
screen "716_TS_IF_NOT_USED" 1280x800, template "Top_Header"
   on GenerateScreen: "SDC_TS_REFERENCE"("SDC\_TS_Nr"); "SDC_TS_IF"(); SetTag("DB_SDC_TS_IF_HMI.HMI[XX].BILD_Nr", 716); SetTag("SDC\_intern_Bildnummer", 716)
   on ClearScreen: SetTag("DB_SDC_TS_IF_HMI.HMI[XX].BILD_Nr", 0)
   TextField "Textfeld_18" at 739,287 size 178x25; Text 'acknowledge error / Command forward'
   Circle "Kreis_27" at 716,292 size 15x15
      Appearance <- "DB_SDC_TS_IF_COMMAND.SEK[XXX].BIT1"
   TextField "Textfeld_1" at 739,304 size 191x25; Text '1 = automatic in section / Command forward'
   Circle "Kreis_1" at 716,308 size 15x15
      Appearance <- "DB_SDC_TS_IF_COMMAND.SEK[XXX].BIT1"
   TextField "Textfeld_2" at 739,319 size 202x25; Text '1 = manual in section / Command forward'
   Circle "Kreis_2" at 716,324 size 15x15
      Appearance <- "DB_SDC_TS_IF_COMMAND.SEK[XXX].BIT1"
   TextField "Textfeld_4" at 739,336 size 201x25; Text 'spare / Command forward / Spare'
   Circle "Kreis_3" at 716,340 size 15x15
      Appearance <- "DB_SDC_TS_IF_COMMAND.SEK[XXX].BIT1"
   TextField "Textfeld_5" at 955,286 size 194x25; Text 'spare / Command forward / Spare'
   Circle "Kreis_4" at 932,291 size 15x15
      Appearance <- "DB_SDC_TS_IF_COMMAND.SEK[XXX].BIT1"
   TextField "Textfeld_6" at 955,303 size 150x25; Text '1 = emergency stop / Command forward'
   Circle "Kreis_5" at 932,307 size 15x15
      Appearance <- "DB_SDC_TS_IF_COMMAND.SEK[XXX].BIT1"
   TextField "Textfeld_7" at 955,318 size 138x25; Text 'spare / Command forward / Spare'
   Circle "Kreis_6" at 932,323 size 15x15
      Appearance <- "DB_SDC_TS_IF_COMMAND.SEK[XXX].BIT1"
   TextField "Textfeld_9" at 738,389 size 125x22; Text 'forward / Command forward'
   Circle "Kreis_8" at 715,394 size 15x15
      Appearance <- "DB_SDC_TS_IF_COMMAND.SEK[XXX].BIT1"
   TextField "Textfeld_10" at 738,406 size 125x22; Text 'backward / Command forward'
   Circle "Kreis_9" at 715,410 size 15x15
      Appearance <- "DB_SDC_TS_IF_COMMAND.SEK[XXX].BIT1"
   TextField "Textfeld_11" at 738,421 size 136x22; Text 'bypass stop position / Command forward'
   Circle "Kreis_10" at 715,426 size 15x15
      Appearance <- "DB_SDC_TS_IF_COMMAND.SEK[XXX].BIT1"
   TextField "Textfeld_12" at 738,438 size 125x22; Text 'speed setpoint 1 / Command forward / Speed Setpoint 1'
   Circle "Kreis_11" at 715,442 size 15x15
      Appearance <- "DB_SDC_TS_IF_COMMAND.SEK[XXX].BIT1"
   TextField "Textfeld_13" at 738,453 size 125x22; Text 'speed setpoint 2 / Command forward / Speed Setpoint 2'
   Circle "Kreis_12" at 715,458 size 15x15
      Appearance <- "DB_SDC_TS_IF_COMMAND.SEK[XXX].BIT1"
   TextField "Textfeld_14" at 738,470 size 156x22; Text 'variable speed setpoint / Command forward / Variable Speed Setpoint'
   Circle "Kreis_13" at 715,474 size 15x15
      Appearance <- "DB_SDC_TS_IF_COMMAND.SEK[XXX].BIT1"
   TextField "Textfeld_15" at 738,485 size 179x22; Text 'enable before stop position / Command forward'
   Circle "Kreis_14" at 715,490 size 15x15
      Appearance <- "DB_SDC_TS_IF_COMMAND.SEK[XXX].BIT1"
   TextField "Textfeld_16" at 738,502 size 168x22; Text 'enable after stop position / Command forward'
   Circle "Kreis_15" at 715,506 size 15x15
      Appearance <- "DB_SDC_TS_IF_COMMAND.SEK[XXX].BIT1"
   TextField "Textfeld_17" at 894,187 size 170x27; Text 'commands / EMS-Number'
   TextField "Textfeld_19" at 625,407 size 27x114; Text 'bits / EMS-Number'
   IOField "EA-Feld_4" at 305,148 size 56x32; FormatPattern 9999
      on OnFinishInput: "SDC_TS_REFERENCE"("SDC\_TS_Nr"); "SDC_TS_IF"()
      ProcessValue <- "SDC\_TS_Nr"
   TextField "Textfeld_3" at 429,151 size 117x23; Text 'section no. / Sektionnumber / Section Number'
   Button "Schaltfläche_1" at 362,148 size 40x32; TextOff '+'
      on Click: function_dd21b452("SDC\_TS_Nr", 1); "SDC_TS_REFERENCE"("SDC\_TS_Nr"); "SDC_TS_IF"()
   Button "Schaltfläche_3" at 265,148 size 39x32; TextOff '-'
      on Click: function_b9b71300("SDC\_TS_Nr", 1); "SDC_TS_REFERENCE"("SDC\_TS_Nr"); "SDC_TS_IF"()
   IOField "EA-Feld_13" at 665,152 size 163x24; Authorization "Benutzerverwaltung"; FormatPattern ????????????????
      Appearance <- "SDC\DB_SDC_TS_PARAMETER\DB_SDC_TS_PARAMETER_HMI.HMI[XX].FR_EDIT"
      ProcessValue <- "SDC\DB_SDC_TS_REFERENCE\DB_SDC_TS_REFERENCE_X.Reference[XXX].Sektion"
      ObjectEnable <- "SDC\DB_SDC_TS_PARAMETER\DB_SDC_TS_PARAMETER_HMI.HMI[XX].FR_EDIT"
   TextField "Textfeld_20" at 625,218 size 27x114; Text 'values / EMS-Number / Values'
   IOField "EA-Feld_1" at 716,221 size 56x28; FormatPattern 99
      on OnFinishInput: "SDC_TS_PARAMETER"(); "SDC_TS_REFERENCE"("SDC\_TS_Nr")
      ProcessValue <- "DB_SDC_TS_IF_COMMAND.SEK[XXX].VAL.PROFIL"
   TextField "Textfeld_21" at 788,223 size 64x25; Text 'car type / Command forward'
   IOField "EA-Feld_2" at 716,237 size 56x28; FormatPattern 999999
      on OnFinishInput: "SDC_TS_PARAMETER"(); "SDC_TS_REFERENCE"("SDC\_TS_Nr")
      ProcessValue <- "DB_SDC_TS_IF_COMMAND.SEK[XXX].VAL.D_SETSPEED"
   TextField "Textfeld_22" at 788,239 size 202x25; Text 'setpoint drive speed mm/min / Command forward'
   IOField "EA-Feld_3" at 716,253 size 56x28; FormatPattern 99999
      on OnFinishInput: "SDC_TS_PARAMETER"(); "SDC_TS_REFERENCE"("SDC\_TS_Nr")
      ProcessValue <- "DB_SDC_TS_IF_COMMAND.SEK[XXX].VAL.D_POS_OFFS"
   TextField "Textfeld_23" at 788,255 size 192x25; Text 'stop position offset mm / Command forward / Stop positions offset mm'
   TextField "Textfeld_24" at 719,369 size 155x22; Text 'drive / Command forward'
   TextField "Textfeld_47" at 738,517 size 166x22; Text 'bypass distance controlle / Command forward / bypass distance control'
   Circle "Kreis_37" at 715,522 size 15x15
      Appearance <- "DB_SDC_TS_IF_COMMAND.SEK[XXX].BIT2"
   TextField "Textfeld_48" at 955,335 size 84x25; Text 'set car type / Command forward'
   Circle "Kreis_38" at 932,339 size 15x15
      Appearance <- "DB_SDC_TS_IF_COMMAND.SEK[XXX].BIT2"
   TextField "Textfeld_49" at 625,657 size 27x59; Text 'fkt / EMS-Number'
   TextField "Textfeld_50" at 766,592 size 155x22; Text 'set / Command forward / Set'
   TextField "Textfeld_51" at 738,612 size 143x22; Text 'EMS to maintenace 1 / Command forward'
   Circle "Kreis_39" at 715,617 size 15x15
      Appearance <- "DB_SDC_TS_IF_COMMAND.SEK[XXX].FKT_SET"
   TextField "Textfeld_52" at 738,629 size 143x22; Text 'EMS to maintenace 2 / Command forward'
   Circle "Kreis_40" at 715,633 size 15x15
      Appearance <- "DB_SDC_TS_IF_COMMAND.SEK[XXX].FKT_SET"
   TextField "Textfeld_53" at 738,644 size 179x22; Text 'emerg. mode without hoist / Command forward'
   Circle "Kreis_41" at 715,649 size 15x15
      Appearance <- "DB_SDC_TS_IF_COMMAND.SEK[XXX].FKT_SET"
   TextField "Textfeld_55" at 738,660 size 129x22; Text 'emerg. mode drive / Command forward'
   Circle "Kreis_43" at 715,665 size 15x15
      Appearance <- "DB_SDC_TS_IF_COMMAND.SEK[XXX].FKT_SET"
   TextField "Textfeld_57" at 738,684 size 125x22; Text 'PE check fault / Command forward / PE Check Fault'
   Circle "Kreis_45" at 715,689 size 15x15
      Appearance <- "DB_SDC_TS_IF_COMMAND.SEK[XXX].FKT_SET"
   TextField "Textfeld_58" at 738,701 size 125x22; Text 'brush check fault / Command forward'
   Circle "Kreis_46" at 715,705 size 15x15
      Appearance <- "DB_SDC_TS_IF_COMMAND.SEK[XXX].FKT_SET"
   TextField "Textfeld_59" at 1054,592 size 155x22; Text 'reset / Command forward / Reset'
   TextField "Textfeld_60" at 1026,612 size 143x22; Text 'EMS to maintenace 1 / Command forward'
   Circle "Kreis_47" at 1003,617 size 15x15
      Appearance <- "DB_SDC_TS_IF_COMMAND.SEK[XXX].FKT_RESET"
   TextField "Textfeld_61" at 1026,629 size 143x22; Text 'EMS to maintenace 2 / Command forward'
   Circle "Kreis_48" at 1003,633 size 15x15
      Appearance <- "DB_SDC_TS_IF_COMMAND.SEK[XXX].FKT_RESET"
   TextField "Textfeld_62" at 1026,644 size 179x22; Text 'emerg. mode without hoist / Command forward'
   Circle "Kreis_49" at 1003,649 size 15x15
      Appearance <- "DB_SDC_TS_IF_COMMAND.SEK[XXX].FKT_RESET"
   TextField "Textfeld_64" at 1026,660 size 129x22; Text 'emerg. mode drive / Command forward'
   Circle "Kreis_51" at 1003,665 size 15x15
      Appearance <- "DB_SDC_TS_IF_COMMAND.SEK[XXX].FKT_RESET"
   TextField "Textfeld_66" at 1026,684 size 125x22; Text 'PE check fault / Command forward / PE Check Fault'
   Circle "Kreis_53" at 1003,689 size 15x15
      Appearance <- "DB_SDC_TS_IF_COMMAND.SEK[XXX].FKT_RESET"
   TextField "Textfeld_67" at 1026,701 size 125x22; Text 'brush check fault / Command forward'
   Circle "Kreis_54" at 1003,705 size 15x15
      Appearance <- "DB_SDC_TS_IF_COMMAND.SEK[XXX].FKT_RESET"
   TextField "Textfeld_68" at 317,193 size 170x27; Text 'status / EMS-Number / Status'
   IOField "EA-Feld_5" at 169,212 size 56x28; FormatPattern 999
      on OnFinishInput: "SDC_TS_PARAMETER"(); "SDC_TS_REFERENCE"("SDC\_TS_Nr")
      ProcessValue <- "DB_SDC_TS_IF_STATUS.SEK[XXX].VAL.EMS_ID"
   TextField "Textfeld_69" at 225,215 size 60x25; Text 'EMS ID / Command forward'
   IOField "EA-Feld_6" at 169,228 size 56x28; FormatPattern 99
      on OnFinishInput: "SDC_TS_PARAMETER"(); "SDC_TS_REFERENCE"("SDC\_TS_Nr")
      ProcessValue <- "DB_SDC_TS_IF_STATUS.SEK[XXX].VAL.PROFIL"
   TextField "Textfeld_70" at 225,231 size 60x25; Text 'car type / Command forward'
   IOField "EA-Feld_7" at 139,244 size 86x28; FormatPattern 9999999999
      on OnFinishInput: "SDC_TS_PARAMETER"(); "SDC_TS_REFERENCE"("SDC\_TS_Nr")
      ProcessValue <- "DB_SDC_TS_IF_STATUS.SEK[XXX].VAL.DRIVE_POS"
   TextField "Textfeld_71" at 225,247 size 170x25; Text 'drive position mm / Command forward'
   IOField "EA-Feld_10" at 385,213 size 56x28; FormatPattern 999
      on OnFinishInput: "SDC_TS_PARAMETER"(); "SDC_TS_REFERENCE"("SDC\_TS_Nr")
      ProcessValue <- "DB_SDC_TS_IF_STATUS.SEK[XXX].VAL.ERROR"
   TextField "Textfeld_74" at 443,215 size 60x25; Text 'error no. / Command forward'
   IOField "EA-Feld_11" at 385,229 size 56x28; FormatPattern 999
      on OnFinishInput: "SDC_TS_PARAMETER"(); "SDC_TS_REFERENCE"("SDC\_TS_Nr")
      ProcessValue <- "DB_SDC_TS_IF_STATUS.SEK[XXX].VAL.DRIVE_POS_PERC"
   TextField "Textfeld_75" at 443,231 size 162x25; Text 'position in % at sektion / Command forward / Position in % in Sektion'
   IOField "EA-Feld_12" at 385,245 size 56x28; FormatPattern 999
      on OnFinishInput: "SDC_TS_PARAMETER"(); "SDC_TS_REFERENCE"("SDC\_TS_Nr")
      ProcessValue <- "DB_SDC_TS_IF_STATUS.SEK[XXX].VAL.SEK"
   TextField "Textfeld_76" at 443,247 size 162x25; Text 'sektion / Command forward / Section'
   TextField "Textfeld_77" at 179,287 size 178x25; Text 'EMS present / Command forward'
   Circle "Kreis_55" at 156,292 size 15x15
      Appearance <- "DB_SDC_TS_IF_STATUS.SEK[XXX].BIT1"
   TextField "Textfeld_78" at 179,304 size 191x25; Text 'general error / Command forward'
   Circle "Kreis_56" at 156,308 size 15x15
      Appearance <- "DB_SDC_TS_IF_STATUS.SEK[XXX].BIT1"
   TextField "Textfeld_79" at 179,319 size 202x25; Text 'EMS in manual mode (IR) / Command forward'
   Circle "Kreis_57" at 156,324 size 15x15
      Appearance <- "DB_SDC_TS_IF_STATUS.SEK[XXX].BIT1"
   TextField "Textfeld_80" at 179,336 size 201x25; Text 'more than 1 EMS in section / Command forward'
   Circle "Kreis_58" at 156,340 size 15x15
      Appearance <- "DB_SDC_TS_IF_STATUS.SEK[XXX].BIT1"
   TextField "Textfeld_81" at 395,286 size 194x25; Text 'error on commands / Command forward'
   Circle "Kreis_59" at 372,291 size 15x15
      Appearance <- "DB_SDC_TS_IF_STATUS.SEK[XXX].BIT1"
   TextField "Textfeld_82" at 395,303 size 229x25; Text 'warning distance controll / Command forward / "1" -> No Stop'
   Circle "Kreis_60" at 372,307 size 15x15
      Appearance <- "DB_SDC_TS_IF_STATUS.SEK[XXX].BIT1"
   TextField "Textfeld_83" at 395,318 size 138x25; Text 'spare / Command forward / Spare'
   Circle "Kreis_61" at 372,323 size 15x15
      Appearance <- "DB_SDC_TS_IF_STATUS.SEK[XXX].BIT1"
   TextField "Textfeld_84" at 395,335 size 220x25; Text 'error code is a warning / Command forward'
   Circle "Kreis_62" at 372,339 size 15x15
      Appearance <- "DB_SDC_TS_IF_STATUS.SEK[XXX].BIT1"
   TextField "Textfeld_85" at 163,369 size 155x22; Text 'drive / Command forward'
   TextField "Textfeld_88" at 186,389 size 125x22; Text 'drive is on / Command forward'
   Circle "Kreis_63" at 163,394 size 15x15
      Appearance <- "DB_SDC_TS_IF_STATUS.SEK[XXX].BIT1"
   TextField "Textfeld_89" at 186,406 size 125x22; Text 'drive is off / Command forward'
   Circle "Kreis_64" at 163,410 size 15x15
      Appearance <- "DB_SDC_TS_IF_STATUS.SEK[XXX].BIT1"
   TextField "Textfeld_94" at 186,421 size 125x22; Text 'in position / Command forward'
   Circle "Kreis_69" at 163,426 size 15x15
      Appearance <- "DB_SDC_TS_IF_STATUS.SEK[XXX].BIT2"
   TextField "Textfeld_95" at 186,437 size 125x22; Text 'before position / Command forward'
   Circle "Kreis_70" at 163,442 size 15x15
      Appearance <- "DB_SDC_TS_IF_STATUS.SEK[XXX].BIT2"
   TextField "Textfeld_96" at 186,453 size 125x22; Text 'after position / Command forward'
   Circle "Kreis_71" at 163,458 size 15x15
      Appearance <- "DB_SDC_TS_IF_STATUS.SEK[XXX].BIT2"
   TextField "Textfeld_97" at 186,469 size 125x22; Text 'after actionpoint 1 / Command forward'
   Circle "Kreis_72" at 163,474 size 15x15
      Appearance <- "DB_SDC_TS_IF_STATUS.SEK[XXX].BIT2"
   TextField "Textfeld_98" at 186,485 size 157x22; Text 'before/at actionpoint 1 / Command forward'
   Circle "Kreis_73" at 163,490 size 15x15
      Appearance <- "DB_SDC_TS_IF_STATUS.SEK[XXX].BIT2"
   TextField "Textfeld_99" at 186,501 size 125x22; Text 'after actionpoint 2 / Command forward'
   Circle "Kreis_74" at 163,506 size 15x15
      Appearance <- "DB_SDC_TS_IF_STATUS.SEK[XXX].BIT2"
   TextField "Textfeld_100" at 186,517 size 152x22; Text 'before/at actionpoint 2 / Command forward'
   Circle "Kreis_75" at 163,522 size 15x15
      Appearance <- "DB_SDC_TS_IF_STATUS.SEK[XXX].BIT2"
   TextField "Textfeld_133" at 186,533 size 125x22; Text 'forwards / Command forward'
   Circle "Kreis_108" at 163,538 size 15x15
      Appearance <- "DB_SDC_TS_IF_STATUS.SEK[XXX].BIT4"
   TextField "Textfeld_134" at 186,550 size 125x22; Text 'backwards / Command forward'
   Circle "Kreis_109" at 163,554 size 15x15
      Appearance <- "DB_SDC_TS_IF_STATUS.SEK[XXX].BIT4"
   TextField "Textfeld_38" at 738,717 size 176x22; Text 'communication check fault / Command forward'
   Circle "Kreis_29" at 715,721 size 15x15
      Appearance <- "DB_SDC_TS_IF_COMMAND.SEK[XXX].FKT_SET"
   TextField "Textfeld_39" at 1026,717 size 176x22; Text 'communication check fault / Command forward'
   Circle "Kreis_30" at 1003,721 size 15x15
      Appearance <- "DB_SDC_TS_IF_COMMAND.SEK[XXX].FKT_RESET"

screen "722_ERRORS_NOT_USED" 1280x800, template "Top_Header"
   on GenerateScreen: "SDC_ERRORS"("HMI_EMS_Nr"); SetTag("SDC\_intern_Bildnummer", 722)
   TextField "Textfeld_18" at 235,235 size 31x132; Text '601 602 603 604 605 606 607 608 Command forward 601'
   Circle "Kreis_27" at 212,238 size 15x15
      Appearance <- "DB_SDC_ERRORS.EMS[XXX].DRIVE_1"
   Circle "Kreis_1" at 212,254 size 15x15
      Appearance <- "DB_SDC_ERRORS.EMS[XXX].DRIVE_1"
   Circle "Kreis_2" at 212,270 size 15x15
      Appearance <- "DB_SDC_ERRORS.EMS[XXX].DRIVE_1"
   Circle "Kreis_3" at 212,286 size 15x15
      Appearance <- "DB_SDC_ERRORS.EMS[XXX].DRIVE_1"
   Circle "Kreis_4" at 212,302 size 15x15
      Appearance <- "DB_SDC_ERRORS.EMS[XXX].DRIVE_1"
   Circle "Kreis_5" at 212,318 size 15x15
      Appearance <- "DB_SDC_ERRORS.EMS[XXX].DRIVE_1"
   Circle "Kreis_6" at 212,334 size 15x15
      Appearance <- "DB_SDC_ERRORS.EMS[XXX].DRIVE_1"
   Circle "Kreis_7" at 212,350 size 15x15
      Appearance <- "DB_SDC_ERRORS.EMS[XXX].DRIVE_1"
   TextField "Textfeld_9" at 292,235 size 31x132; Text '609 610 611 612 613 614 615 616 Command forward 609'
   Circle "Kreis_8" at 269,238 size 15x15
      Appearance <- "DB_SDC_ERRORS.EMS[XXX].DRIVE_1"
   Circle "Kreis_9" at 269,254 size 15x15
      Appearance <- "DB_SDC_ERRORS.EMS[XXX].DRIVE_1"
   Circle "Kreis_10" at 269,270 size 15x15
      Appearance <- "DB_SDC_ERRORS.EMS[XXX].DRIVE_1"
   Circle "Kreis_11" at 269,286 size 15x15
      Appearance <- "DB_SDC_ERRORS.EMS[XXX].DRIVE_1"
   Circle "Kreis_12" at 269,302 size 15x15
      Appearance <- "DB_SDC_ERRORS.EMS[XXX].DRIVE_1"
   Circle "Kreis_13" at 269,318 size 15x15
      Appearance <- "DB_SDC_ERRORS.EMS[XXX].DRIVE_1"
   Circle "Kreis_14" at 269,334 size 15x15
      Appearance <- "DB_SDC_ERRORS.EMS[XXX].DRIVE_1"
   Circle "Kreis_15" at 269,350 size 15x15
      Appearance <- "DB_SDC_ERRORS.EMS[XXX].DRIVE_1"
   TextField "Textfeld_17" at 271,202 size 100x38; Text 'drive / EMS-Number / Drive'
   TextField "Textfeld_19" at 180,241 size 32x114; Text 'generally / EMS-Number / General'
   IOField "EA-Feld_4" at 265,156 size 56x32; FormatPattern 9999
      on OnFinishInput: "SDC_EMS_STATUS"("HMI_EMS_Nr"); "SDC_TS_REFERENCE"("SDC\DB_SDC_EMS\EMS[XXX].TS_STAT.VAL.SEK"); "SDC_EMS_TA_STATUS"("HMI_EMS_Nr"); "SDC_ERRORS"("HMI_EMS_Nr"); SetTag("_DB_SDC_ERRORS.Error_nr", "SDC\DB_SDC_EMS\EMS[XXX].TS_STAT.VAL.ERROR")
      ProcessValue <- "HMI_EMS_Nr"
   Button "Schaltfläche_1" at 322,156 size 40x32; TextOff '+'
      on Click: function_dd21b452("HMI_EMS_Nr", 1); "SDC_EMS_STATUS"("HMI_EMS_Nr"); "SDC_TS_REFERENCE"("SDC\DB_SDC_EMS\EMS[XXX].TS_STAT.VAL.SEK"); "SDC_EMS_TA_STATUS"("HMI_EMS_Nr"); "SDC_ERRORS"("HMI_EMS_Nr"); SetTag("_DB_SDC_ERRORS.Error_nr", "SDC\DB_SDC_EMS\EMS[XXX].TS_STAT.VAL.ERROR")
   Button "Schaltfläche_3" at 225,156 size 39x32; TextOff '-'
      on Click: function_b9b71300("HMI_EMS_Nr", 1); "SDC_EMS_STATUS"("HMI_EMS_Nr"); "SDC_TS_REFERENCE"("SDC\DB_SDC_EMS\EMS[XXX].TS_STAT.VAL.SEK"); "SDC_EMS_TA_STATUS"("HMI_EMS_Nr"); "SDC_ERRORS"("HMI_EMS_Nr"); SetTag("_DB_SDC_ERRORS.Error_nr", "SDC\DB_SDC_EMS\EMS[XXX].TS_STAT.VAL.ERROR")
   TextField "Textfeld_3" at 373,159 size 102x23; Text 'EMS-No. / EMS-Number / EMS-Nummer'
   TextField "Textfeld_20" at 235,371 size 31x132; Text '633 634 635 636 637 638 639 640 Command forward 633'
   Circle "Kreis_16" at 212,374 size 15x15
      Appearance <- "DB_SDC_ERRORS.EMS[XXX].FC_DRIVE_1"
   Circle "Kreis_17" at 212,390 size 15x15
      Appearance <- "DB_SDC_ERRORS.EMS[XXX].FC_DRIVE_1"
   Circle "Kreis_18" at 212,406 size 15x15
      Appearance <- "DB_SDC_ERRORS.EMS[XXX].FC_DRIVE_1"
   Circle "Kreis_19" at 212,422 size 15x15
      Appearance <- "DB_SDC_ERRORS.EMS[XXX].FC_DRIVE_1"
   Circle "Kreis_20" at 212,438 size 15x15
      Appearance <- "DB_SDC_ERRORS.EMS[XXX].FC_DRIVE_1"
   Circle "Kreis_21" at 212,454 size 15x15
      Appearance <- "DB_SDC_ERRORS.EMS[XXX].FC_DRIVE_1"
   Circle "Kreis_22" at 212,470 size 15x15
      Appearance <- "DB_SDC_ERRORS.EMS[XXX].FC_DRIVE_1"
   Circle "Kreis_23" at 212,486 size 15x15
      Appearance <- "DB_SDC_ERRORS.EMS[XXX].FC_DRIVE_1"
   TextField "Textfeld_28" at 292,371 size 31x132; Text '641 642 643 644 645 646 647 648 Command forward 641'
   Circle "Kreis_24" at 269,374 size 15x15
      Appearance <- "DB_SDC_ERRORS.EMS[XXX].FC_DRIVE_1"
   Circle "Kreis_25" at 269,390 size 15x15
      Appearance <- "DB_SDC_ERRORS.EMS[XXX].FC_DRIVE_1"
   Circle "Kreis_26" at 269,406 size 15x15
      Appearance <- "DB_SDC_ERRORS.EMS[XXX].FC_DRIVE_1"
   Circle "Kreis_28" at 269,422 size 15x15
      Appearance <- "DB_SDC_ERRORS.EMS[XXX].FC_DRIVE_1"
   Circle "Kreis_29" at 269,438 size 15x15
      Appearance <- "DB_SDC_ERRORS.EMS[XXX].FC_DRIVE_1"
   Circle "Kreis_30" at 269,454 size 15x15
      Appearance <- "DB_SDC_ERRORS.EMS[XXX].FC_DRIVE_1"
   Circle "Kreis_31" at 269,470 size 15x15
      Appearance <- "DB_SDC_ERRORS.EMS[XXX].FC_DRIVE_1"
   Circle "Kreis_32" at 269,486 size 15x15
      Appearance <- "DB_SDC_ERRORS.EMS[XXX].FC_DRIVE_1"
   TextField "Textfeld_36" at 167,377 size 32x119; Text 'FC / EMS-Number / Frequency Conv'
   TextField "Textfeld_37" at 235,507 size 31x132; Text '649 650 651 652 653 654 655 656 Command forward 649'
   Circle "Kreis_33" at 212,510 size 15x15
      Appearance <- "DB_SDC_ERRORS.EMS[XXX].SAFETY_DRIVE"
   Circle "Kreis_34" at 212,526 size 15x15
      Appearance <- "DB_SDC_ERRORS.EMS[XXX].SAFETY_DRIVE"
   Circle "Kreis_35" at 212,542 size 15x15
      Appearance <- "DB_SDC_ERRORS.EMS[XXX].SAFETY_DRIVE"
   Circle "Kreis_36" at 212,558 size 15x15
      Appearance <- "DB_SDC_ERRORS.EMS[XXX].SAFETY_DRIVE"
   Circle "Kreis_37" at 212,574 size 15x15
      Appearance <- "DB_SDC_ERRORS.EMS[XXX].SAFETY_DRIVE"
   Circle "Kreis_38" at 212,590 size 15x15
      Appearance <- "DB_SDC_ERRORS.EMS[XXX].SAFETY_DRIVE"
   Circle "Kreis_39" at 212,606 size 15x15
      Appearance <- "DB_SDC_ERRORS.EMS[XXX].SAFETY_DRIVE"
   Circle "Kreis_40" at 212,622 size 15x15
      Appearance <- "DB_SDC_ERRORS.EMS[XXX].SAFETY_DRIVE"
   TextField "Textfeld_45" at 292,507 size 31x132; Text '657 658 659 660 661 662 663 664 Command forward 657'
   Circle "Kreis_41" at 269,510 size 15x15
      Appearance <- "DB_SDC_ERRORS.EMS[XXX].SAFETY_DRIVE"
   Circle "Kreis_42" at 269,526 size 15x15
      Appearance <- "DB_SDC_ERRORS.EMS[XXX].SAFETY_DRIVE"
   Circle "Kreis_43" at 269,542 size 15x15
      Appearance <- "DB_SDC_ERRORS.EMS[XXX].SAFETY_DRIVE"
   Circle "Kreis_44" at 269,558 size 15x15
      Appearance <- "DB_SDC_ERRORS.EMS[XXX].SAFETY_DRIVE"
   Circle "Kreis_45" at 269,574 size 15x15
      Appearance <- "DB_SDC_ERRORS.EMS[XXX].SAFETY_DRIVE"
   Circle "Kreis_46" at 269,590 size 15x15
      Appearance <- "DB_SDC_ERRORS.EMS[XXX].SAFETY_DRIVE"
   Circle "Kreis_47" at 269,606 size 15x15
      Appearance <- "DB_SDC_ERRORS.EMS[XXX].SAFETY_DRIVE"
   Circle "Kreis_48" at 269,622 size 15x15
      Appearance <- "DB_SDC_ERRORS.EMS[XXX].SAFETY_DRIVE"
   TextField "Textfeld_53" at 180,511 size 32x76; Text 'safety / EMS-Number / Safety'
   TextField "Textfeld_54" at 355,235 size 31x132; Text '617 618 619 620 621 622 623 624 Command forward 617'
   Circle "Kreis_49" at 332,238 size 15x15
      Appearance <- "DB_SDC_ERRORS.EMS[XXX].DRIVE_2"
   Circle "Kreis_50" at 332,254 size 15x15
      Appearance <- "DB_SDC_ERRORS.EMS[XXX].DRIVE_2"
   Circle "Kreis_51" at 332,270 size 15x15
      Appearance <- "DB_SDC_ERRORS.EMS[XXX].DRIVE_2"
   Circle "Kreis_52" at 332,286 size 15x15
      Appearance <- "DB_SDC_ERRORS.EMS[XXX].DRIVE_2"
   Circle "Kreis_53" at 332,302 size 15x15
      Appearance <- "DB_SDC_ERRORS.EMS[XXX].DRIVE_2"
   Circle "Kreis_54" at 332,318 size 15x15
      Appearance <- "DB_SDC_ERRORS.EMS[XXX].DRIVE_2"
   Circle "Kreis_55" at 332,334 size 15x15
      Appearance <- "DB_SDC_ERRORS.EMS[XXX].DRIVE_2"
   Circle "Kreis_56" at 332,350 size 15x15
      Appearance <- "DB_SDC_ERRORS.EMS[XXX].DRIVE_2"
   TextField "Textfeld_62" at 412,235 size 31x132; Text '625 626 627 628 629 630 631 632 Command forward 625'
   Circle "Kreis_57" at 389,238 size 15x15
      Appearance <- "DB_SDC_ERRORS.EMS[XXX].DRIVE_2"
   Circle "Kreis_58" at 389,254 size 15x15
      Appearance <- "DB_SDC_ERRORS.EMS[XXX].DRIVE_2"
   Circle "Kreis_59" at 389,270 size 15x15
      Appearance <- "DB_SDC_ERRORS.EMS[XXX].DRIVE_2"
   Circle "Kreis_60" at 389,286 size 15x15
      Appearance <- "DB_SDC_ERRORS.EMS[XXX].DRIVE_2"
   Circle "Kreis_61" at 389,302 size 15x15
      Appearance <- "DB_SDC_ERRORS.EMS[XXX].DRIVE_2"
   Circle "Kreis_62" at 389,318 size 15x15
      Appearance <- "DB_SDC_ERRORS.EMS[XXX].DRIVE_2"
   Circle "Kreis_63" at 389,334 size 15x15
      Appearance <- "DB_SDC_ERRORS.EMS[XXX].DRIVE_2"
   Circle "Kreis_64" at 389,350 size 15x15
      Appearance <- "DB_SDC_ERRORS.EMS[XXX].DRIVE_2"
   TextField "Textfeld_70" at 355,371 size 31x132; Text '665 666 667 668 669 670 671 672 Command forward 665'
   Circle "Kreis_65" at 332,374 size 15x15
      Appearance <- "DB_SDC_ERRORS.EMS[XXX].FC_DRIVE_2"
   Circle "Kreis_66" at 332,390 size 15x15
      Appearance <- "DB_SDC_ERRORS.EMS[XXX].FC_DRIVE_2"
   Circle "Kreis_67" at 332,406 size 15x15
      Appearance <- "DB_SDC_ERRORS.EMS[XXX].FC_DRIVE_2"
   Circle "Kreis_68" at 332,422 size 15x15
      Appearance <- "DB_SDC_ERRORS.EMS[XXX].FC_DRIVE_2"
   Circle "Kreis_69" at 332,438 size 15x15
      Appearance <- "DB_SDC_ERRORS.EMS[XXX].FC_DRIVE_2"
   Circle "Kreis_70" at 332,454 size 15x15
      Appearance <- "DB_SDC_ERRORS.EMS[XXX].FC_DRIVE_2"
   Circle "Kreis_71" at 332,470 size 15x15
      Appearance <- "DB_SDC_ERRORS.EMS[XXX].FC_DRIVE_2"
   Circle "Kreis_72" at 332,486 size 15x15
      Appearance <- "DB_SDC_ERRORS.EMS[XXX].FC_DRIVE_2"
   TextField "Textfeld_78" at 412,371 size 31x132; Text '673 674 675 676 677 678 679 680 Command forward 673'
   Circle "Kreis_73" at 389,374 size 15x15
      Appearance <- "DB_SDC_ERRORS.EMS[XXX].FC_DRIVE_2"
   Circle "Kreis_74" at 389,390 size 15x15
      Appearance <- "DB_SDC_ERRORS.EMS[XXX].FC_DRIVE_2"
   Circle "Kreis_75" at 389,406 size 15x15
      Appearance <- "DB_SDC_ERRORS.EMS[XXX].FC_DRIVE_2"
   Circle "Kreis_76" at 389,422 size 15x15
      Appearance <- "DB_SDC_ERRORS.EMS[XXX].FC_DRIVE_2"
   Circle "Kreis_77" at 389,438 size 15x15
      Appearance <- "DB_SDC_ERRORS.EMS[XXX].FC_DRIVE_2"
   Circle "Kreis_78" at 389,454 size 15x15
      Appearance <- "DB_SDC_ERRORS.EMS[XXX].FC_DRIVE_2"
   Circle "Kreis_79" at 389,470 size 15x15
      Appearance <- "DB_SDC_ERRORS.EMS[XXX].FC_DRIVE_2"
   Circle "Kreis_80" at 389,486 size 15x15
      Appearance <- "DB_SDC_ERRORS.EMS[XXX].FC_DRIVE_2"
   TextField "Textfeld_86" at 483,235 size 31x132; Text '701 702 703 704 705 706 707 708 Command forward 701'
   Circle "Kreis_81" at 460,238 size 15x15
      Appearance <- "DB_SDC_ERRORS.EMS[XXX].HOIST_1"
   Circle "Kreis_82" at 460,254 size 15x15
      Appearance <- "DB_SDC_ERRORS.EMS[XXX].HOIST_1"
   Circle "Kreis_83" at 460,270 size 15x15
      Appearance <- "DB_SDC_ERRORS.EMS[XXX].HOIST_1"
   Circle "Kreis_84" at 460,286 size 15x15
      Appearance <- "DB_SDC_ERRORS.EMS[XXX].HOIST_1"
   Circle "Kreis_85" at 460,302 size 15x15
      Appearance <- "DB_SDC_ERRORS.EMS[XXX].HOIST_1"
   Circle "Kreis_86" at 460,318 size 15x15
      Appearance <- "DB_SDC_ERRORS.EMS[XXX].HOIST_1"
   Circle "Kreis_87" at 460,334 size 15x15
      Appearance <- "DB_SDC_ERRORS.EMS[XXX].HOIST_1"
   Circle "Kreis_88" at 460,350 size 15x15
      Appearance <- "DB_SDC_ERRORS.EMS[XXX].HOIST_1"
   TextField "Textfeld_94" at 540,235 size 31x132; Text '709 710 711 712 713 714 715 716 Command forward 709'
   Circle "Kreis_89" at 517,238 size 15x15
      Appearance <- "DB_SDC_ERRORS.EMS[XXX].HOIST_1"
   Circle "Kreis_90" at 517,254 size 15x15
      Appearance <- "DB_SDC_ERRORS.EMS[XXX].HOIST_1"
   Circle "Kreis_91" at 517,270 size 15x15
      Appearance <- "DB_SDC_ERRORS.EMS[XXX].HOIST_1"
   Circle "Kreis_92" at 517,286 size 15x15
      Appearance <- "DB_SDC_ERRORS.EMS[XXX].HOIST_1"
   Circle "Kreis_93" at 517,302 size 15x15
      Appearance <- "DB_SDC_ERRORS.EMS[XXX].HOIST_1"
   Circle "Kreis_94" at 517,318 size 15x15
      Appearance <- "DB_SDC_ERRORS.EMS[XXX].HOIST_1"
   Circle "Kreis_95" at 517,334 size 15x15
      Appearance <- "DB_SDC_ERRORS.EMS[XXX].HOIST_1"
   Circle "Kreis_96" at 517,350 size 15x15
      Appearance <- "DB_SDC_ERRORS.EMS[XXX].HOIST_1"
   TextField "Textfeld_102" at 516,202 size 100x38; Text 'hoist / EMS-Number / Hoist'
   TextField "Textfeld_104" at 483,371 size 31x132; Text '733 734 735 736 737 738 739 740 Command forward 733'
   Circle "Kreis_97" at 460,374 size 15x15
      Appearance <- "DB_SDC_ERRORS.EMS[XXX].FC_HOIST_1"
   Circle "Kreis_98" at 460,390 size 15x15
      Appearance <- "DB_SDC_ERRORS.EMS[XXX].FC_HOIST_1"
   Circle "Kreis_99" at 460,406 size 15x15
      Appearance <- "DB_SDC_ERRORS.EMS[XXX].FC_HOIST_1"
   Circle "Kreis_100" at 460,422 size 15x15
      Appearance <- "DB_SDC_ERRORS.EMS[XXX].FC_HOIST_1"
   Circle "Kreis_101" at 460,438 size 15x15
      Appearance <- "DB_SDC_ERRORS.EMS[XXX].FC_HOIST_1"
   Circle "Kreis_102" at 460,454 size 15x15
      Appearance <- "DB_SDC_ERRORS.EMS[XXX].FC_HOIST_1"
   Circle "Kreis_103" at 460,470 size 15x15
      Appearance <- "DB_SDC_ERRORS.EMS[XXX].FC_HOIST_1"
   Circle "Kreis_104" at 460,486 size 15x15
      Appearance <- "DB_SDC_ERRORS.EMS[XXX].FC_HOIST_1"
   TextField "Textfeld_112" at 540,371 size 31x132; Text '741 742 743 744 745 746 747 748 Command forward 741'
   Circle "Kreis_105" at 517,374 size 15x15
      Appearance <- "DB_SDC_ERRORS.EMS[XXX].FC_HOIST_1"
   Circle "Kreis_106" at 517,390 size 15x15
      Appearance <- "DB_SDC_ERRORS.EMS[XXX].FC_HOIST_1"
   Circle "Kreis_107" at 517,406 size 15x15
      Appearance <- "DB_SDC_ERRORS.EMS[XXX].FC_HOIST_1"
   Circle "Kreis_108" at 517,422 size 15x15
      Appearance <- "DB_SDC_ERRORS.EMS[XXX].FC_HOIST_1"
   Circle "Kreis_109" at 517,438 size 15x15
      Appearance <- "DB_SDC_ERRORS.EMS[XXX].FC_HOIST_1"
   Circle "Kreis_110" at 517,454 size 15x15
      Appearance <- "DB_SDC_ERRORS.EMS[XXX].FC_HOIST_1"
   Circle "Kreis_111" at 517,470 size 15x15
      Appearance <- "DB_SDC_ERRORS.EMS[XXX].FC_HOIST_1"
   Circle "Kreis_112" at 517,486 size 15x15
      Appearance <- "DB_SDC_ERRORS.EMS[XXX].FC_HOIST_1"
   TextField "Textfeld_121" at 483,507 size 31x132; Text '749 750 751 752 753 754 755 756 Command forward 749'
   Circle "Kreis_113" at 460,510 size 15x15
      Appearance <- "DB_SDC_ERRORS.EMS[XXX].SAFETY_HOIST"
   Circle "Kreis_114" at 460,526 size 15x15
      Appearance <- "DB_SDC_ERRORS.EMS[XXX].SAFETY_HOIST"
   Circle "Kreis_115" at 460,542 size 15x15
      Appearance <- "DB_SDC_ERRORS.EMS[XXX].SAFETY_HOIST"
   Circle "Kreis_116" at 460,558 size 15x15
      Appearance <- "DB_SDC_ERRORS.EMS[XXX].SAFETY_HOIST"
   Circle "Kreis_117" at 460,574 size 15x15
      Appearance <- "DB_SDC_ERRORS.EMS[XXX].SAFETY_HOIST"
   Circle "Kreis_118" at 460,590 size 15x15
      Appearance <- "DB_SDC_ERRORS.EMS[XXX].SAFETY_HOIST"
   Circle "Kreis_119" at 460,606 size 15x15
      Appearance <- "DB_SDC_ERRORS.EMS[XXX].SAFETY_HOIST"
   Circle "Kreis_120" at 460,622 size 15x15
      Appearance <- "DB_SDC_ERRORS.EMS[XXX].SAFETY_HOIST"
   TextField "Textfeld_129" at 540,507 size 31x132; Text '757 758 759 760 761 762 763 764 Command forward 757'
   Circle "Kreis_121" at 517,510 size 15x15
      Appearance <- "DB_SDC_ERRORS.EMS[XXX].SAFETY_HOIST"
   Circle "Kreis_122" at 517,526 size 15x15
      Appearance <- "DB_SDC_ERRORS.EMS[XXX].SAFETY_HOIST"
   Circle "Kreis_123" at 517,542 size 15x15
      Appearance <- "DB_SDC_ERRORS.EMS[XXX].SAFETY_HOIST"
   Circle "Kreis_124" at 517,558 size 15x15
      Appearance <- "DB_SDC_ERRORS.EMS[XXX].SAFETY_HOIST"
   Circle "Kreis_125" at 517,574 size 15x15
      Appearance <- "DB_SDC_ERRORS.EMS[XXX].SAFETY_HOIST"
   Circle "Kreis_126" at 517,590 size 15x15
      Appearance <- "DB_SDC_ERRORS.EMS[XXX].SAFETY_HOIST"
   Circle "Kreis_127" at 517,606 size 15x15
      Appearance <- "DB_SDC_ERRORS.EMS[XXX].SAFETY_HOIST"
   Circle "Kreis_128" at 517,622 size 15x15
      Appearance <- "DB_SDC_ERRORS.EMS[XXX].SAFETY_HOIST"
   TextField "Textfeld_138" at 603,235 size 31x132; Text '717 718 719 720 721 722 723 724 Command forward 717'
   Circle "Kreis_129" at 580,238 size 15x15
      Appearance <- "DB_SDC_ERRORS.EMS[XXX].HOIST_2"
   Circle "Kreis_130" at 580,254 size 15x15
      Appearance <- "DB_SDC_ERRORS.EMS[XXX].HOIST_2"
   Circle "Kreis_131" at 580,270 size 15x15
      Appearance <- "DB_SDC_ERRORS.EMS[XXX].HOIST_2"
   Circle "Kreis_132" at 580,286 size 15x15
      Appearance <- "DB_SDC_ERRORS.EMS[XXX].HOIST_2"
   Circle "Kreis_133" at 580,302 size 15x15
      Appearance <- "DB_SDC_ERRORS.EMS[XXX].HOIST_2"
   Circle "Kreis_134" at 580,318 size 15x15
      Appearance <- "DB_SDC_ERRORS.EMS[XXX].HOIST_2"
   Circle "Kreis_135" at 580,334 size 15x15
      Appearance <- "DB_SDC_ERRORS.EMS[XXX].HOIST_2"
   Circle "Kreis_136" at 580,350 size 15x15
      Appearance <- "DB_SDC_ERRORS.EMS[XXX].HOIST_2"
   TextField "Textfeld_146" at 660,235 size 31x132; Text '725 726 727 728 729 730 731 732 Command forward 725'
   Circle "Kreis_137" at 637,238 size 15x15
      Appearance <- "DB_SDC_ERRORS.EMS[XXX].HOIST_2"
   Circle "Kreis_138" at 637,254 size 15x15
      Appearance <- "DB_SDC_ERRORS.EMS[XXX].HOIST_2"
   Circle "Kreis_139" at 637,270 size 15x15
      Appearance <- "DB_SDC_ERRORS.EMS[XXX].HOIST_2"
   Circle "Kreis_140" at 637,286 size 15x15
      Appearance <- "DB_SDC_ERRORS.EMS[XXX].HOIST_2"
   Circle "Kreis_141" at 637,302 size 15x15
      Appearance <- "DB_SDC_ERRORS.EMS[XXX].HOIST_2"
   Circle "Kreis_142" at 637,318 size 15x15
      Appearance <- "DB_SDC_ERRORS.EMS[XXX].HOIST_2"
   Circle "Kreis_143" at 637,334 size 15x15
      Appearance <- "DB_SDC_ERRORS.EMS[XXX].HOIST_2"
   Circle "Kreis_144" at 637,350 size 15x15
      Appearance <- "DB_SDC_ERRORS.EMS[XXX].HOIST_2"
   TextField "Textfeld_154" at 603,371 size 31x132; Text '765 766 767 768 769 770 771 772 Command forward 765'
   Circle "Kreis_145" at 580,374 size 15x15
      Appearance <- "DB_SDC_ERRORS.EMS[XXX].FC_HOIST_2"
   Circle "Kreis_146" at 580,390 size 15x15
      Appearance <- "DB_SDC_ERRORS.EMS[XXX].FC_HOIST_2"
   Circle "Kreis_147" at 580,406 size 15x15
      Appearance <- "DB_SDC_ERRORS.EMS[XXX].FC_HOIST_2"
   Circle "Kreis_148" at 580,422 size 15x15
      Appearance <- "DB_SDC_ERRORS.EMS[XXX].FC_HOIST_2"
   Circle "Kreis_149" at 580,438 size 15x15
      Appearance <- "DB_SDC_ERRORS.EMS[XXX].FC_HOIST_2"
   Circle "Kreis_150" at 580,454 size 15x15
      Appearance <- "DB_SDC_ERRORS.EMS[XXX].FC_HOIST_2"
   Circle "Kreis_151" at 580,470 size 15x15
      Appearance <- "DB_SDC_ERRORS.EMS[XXX].FC_HOIST_2"
   Circle "Kreis_152" at 580,486 size 15x15
      Appearance <- "DB_SDC_ERRORS.EMS[XXX].FC_HOIST_2"
   TextField "Textfeld_162" at 660,371 size 31x132; Text '773 774 775 776 777 778 779 780 Command forward 773'
   Circle "Kreis_153" at 637,374 size 15x15
      Appearance <- "DB_SDC_ERRORS.EMS[XXX].FC_HOIST_2"
   Circle "Kreis_154" at 637,390 size 15x15
      Appearance <- "DB_SDC_ERRORS.EMS[XXX].FC_HOIST_2"
   Circle "Kreis_155" at 637,406 size 15x15
      Appearance <- "DB_SDC_ERRORS.EMS[XXX].FC_HOIST_2"
   Circle "Kreis_156" at 637,422 size 15x15
      Appearance <- "DB_SDC_ERRORS.EMS[XXX].FC_HOIST_2"